        [0].6   // Pylon Home Sensor/Encoder Incongruence - -B26002I -B26007I
        [0].7   // Pylon Home Sensor/Encoder Incongruence - -B26002I -B26007I
        [2].30   // Code 2.30 Pylon Angle overlimit Alarm by Encoder
        [2].16   // Code 2.16 DC Converter Mot 1_3 Rif. T608C DRIVE FAULT
        [0].2   // Gondola Motor 5 Overvoltage Ref. K706C
        [0].10   // Compressor Motor Protection Feedback -F18002C
        [0].0   // Motor 1 Overvoltage control - Relay OK -K10302G
        [1].0   // Gondola Communication Modem Fault CH1 & CH2 -T27002C
        [0].11   // Motor 5 Overvoltage control - Relay OK -K14302G
        [1].1   // Code 1.1 Contactor QC8201H Fault feedback OFF status
        [1].3   // Code 1.3 Contactor QC8204H Fault feedback OFF status
        [0].12   // Motor 6 Overvoltage control - Relay OK -K14307G
        [0].1   // Motor 2 Overvoltage control - Relay OK -K10307G
        [1].5   // Code 1.5 Contactor QC8206H Fault feedback OFF status
        [1].2   // Code 1.2 Contactor QC8201H Fault feedback ON status
        [0].3   // Motor 3 Overvoltage control - Relay OK -K12302G
        [1].4   // Code 1.4 Contactor QC8204H Fault feedback ON status
        [0].4   // Motor 4 Overvoltage control - Relay OK -K12307G
        [1].6   // Code 1.6 Contactor QC8206H Fault feedback ON status
        [1].7   // Pylon Motor 2/4 Fault
        [1].8   // Pylon Motor 1/3 Fault
   Emergencies_Std_CL1 : DINT[8];
        [1].0   // Motor 1-2 Fan Protection Feedback -F10402C -F10406C
        [1].2   // Motor 3-4 Fan Protection Feedback -F12402C -F12406C
        [1].11   // Motor 5 Thermal Probe -K14702H
        [1].3   // Motor 5-6 Fan Protection Feedback -F14402C -F14406C
        [1].12   // Motor 4 Thermal Probe -K12704H
        [1].13   // Motor 6 Thermal Probe -K14704H
        [2].0   // Module K20510C Fault
        [2].1   // Module K20511C Fault
        [2].2   // Module K20512C Fault
        [2].3   // Module K20513C Fault
        [2].4   // Module K20514C Fault
        [2].5   // Module K20515C Fault
        [2].6   // Module K20516C Fault
        [2].7   // Module K20517C Fault
        [1].14   // Motor 7 Thermal Probe -K16602H
        [1].1   // Motor 7 Fan Protection Feedback -F16402C
        [1].6   // MCC High temeprature -S75003C
        [1].8   // Motor 1 Thermal Probe -K10702H
        [1].9   // Motor 2 Thermal Probe -K10704H
        [1].4   // Gondola Motor 7 Fault
        [1].5   // Pylon Motor 5/6 Fault
   Emergency_Brake_manual_Cmd : BOOL;
   Emergency_Brake_manual_Perm : BOOL := 1;
   Emergency_Brake_SL : ALIAS FOR K300_OCC:6:O.6;   // _S31207D
   Emergency_Captr : DINT[11] := ([0] := 1024, [1] := 384, [2] := 1062171331, [4] := 1062171331);
   Enable_to_Start : UDT_CROUT := (CROUT.Feedback1 := 1, CROUT.Feedback2 := 1, CROUT.InputStatus := 1, CROUT.OutputStatus := 1, CROUT.FeedbackReactionTime := 200, Out_Status := 1);   // Abilitazione allo start QC8011E QC8013E
   Encoder_Resetted : BOOL;
   Fault_2_4 : Powerflex_DC_Fault := (Fault_Code := 75);
   Fault_7 : Powerflex_DC_Fault := (Fault_Code := 75);
   FeedBack_Drives_Contactors : BOOL := 1;
   First_Push_Set_Torque_to_Zero : BOOL;
   Flyng_Start_Req : BOOL;
   Gate_Entry_Unlock_Selector : BOOL := 1;   // -S30701F
   Gate_Exit_Unlock_Selector : BOOL := 1;   // -S30705F
   Gate_Magnalock_Enable : UDT_CROUT := (CROUT.Actuate := 1, CROUT.InputStatus := 1, CROUT.OutputStatus := 1, CROUT.FeedbackReactionTime := 250, CROUT.FP := 1, CROUT.FaultCode := 20483);   // Gate Lock Enable -Q25102E
   Gate_Operator_Unlock_Selector : BOOL;   // -S30707F
   GateCommand : DINT := 416;
        .5   // Gate 1 Open
        .7   // Gate 2 Open
        .9   // Gate 3 Open
        .4   // Gate 1 Close
        .6   // Gate 2 Close
        .8   // Gate 3 Close
   GateRequest : DINT;
        .5   // Gate 1 Open
        .7   // Gate 2 Open
        .9   // Gate 3 Open
        .4   // Gate 1 Close
        .6   // Gate 2 Close
        .8   // Gate 3 Close
   Gates_Auto_Release : BOOL;   // .. At end of Cycle Open Gates Open RESTRAINTS
   Gates_Open_Permissive : Permissive := (All_Permissive_Ok := 1, BitsConditions := -1);
   Girella_Field_Actuate_During_Inactivity : BOOL;
   Girella_Gradi_Sec : DINT := 20;
   Gondola_Axe : Axe := (Speed := -5.538001e-24, Speed_ABS := 5.538001e-24);
   Gondola_Decc_timer_Start : BOOL;
   Gondola_Direction_CW_1 : BOOL;   // 0 > CCW 1 > CW
   Gondola_Direction_CW_2 : BOOL := 1;   // 0 > CCW 1 > CW
   Gondola_Drive_Enable : UDT_CROUT := (CROUT.Feedback1 := 1, CROUT.Feedback2 := 1, CROUT.InputStatus := 1, CROUT.OutputStatus := 1, CROUT.FeedbackReactionTime := 1000);   // Gondola Drive Ch1-Ch2 Start Enable Contactors -Q16105E -Q16107E
   Gondola_Immediatly_Stop : BOOL := 1;
   Gondola_Out_Ref : INT;
   Gondola_Speed_Ref_ABS : REAL;
   Gondola_Speed_Reference : DINT;
   Gondola_Standstill_from_inertia : BOOL := 1;
   Gondola_Stop_Beginning : BOOL;
   Gondola_Stop_CW : BOOL := 1;   // Gondola Sto Direction 0 > CCW 1 > CW
   Gondola_Stop_IP : BOOL;   // Gondola Stop Sequence In Progress
   Gondola_Stop_Step : DINT;
   Gondola_Torque_Lim : REAL := 100.0;
   HLL_T1_R011 : HL_LIMIT := (HighLimit := 77.39982, LowLimit := -77.39982);
   HMI_Angle : REAL;
   HMI_Auto_Cycle_in_Modify : Auto_Cycle := (Pylon_Angle := 120, Cycle_Time_min := 2, Cycle_Time_sec := 25, Gondola_Speed[0] := 20, Gondola_Speed[1] := 70, Gondola_Speed[2] := -75, Gondola_Speed[3] := 50, Gondola_Time[1] := 60, Gondola_Time[2] := 50, Gondola_Time[3] := 20);
   HMI_Auto_Cycle_Step_Modify : DINT := 2;
   HMI_button_addtoindex : BOOL;
   HMI_button_subtracttoindex : BOOL;
   HMI_Current_Screen : DINT;
   HMI_Disable_external_acces : BOOL;   // ROUTER A72A07D Disable external acces
   HMI_Drive_Fault_Descr : STRING[4] := ([1] := 'Communication card fault Port 5', [2] := 'Pommunication card fault Port 5', [3] := 'Pommunication card fault Port 5');
        [0]   // Pylon motor 1 3
        [1]   // Pylon motor 2 4
        [2]   // Gondola motor 5
   HMI_Enable_external_acces : BOOL;   // ROUTER A72A07D Eneble external acces
   HMI_Gondola_Start_Delay : DINT := 5;
   HMI_Horn_Pb : BOOL;   // HMIN Horn Pushbutton
   HMI_JM_Stats_Hist : Run_Count_Hist_JM[10];
   HMI_Lamp_Test : BOOL;
   HMI_Light_Pb : BOOL;
   HMI_Modify_Auto_Cycle_Ptr : DINT := 1;
   HMI_Monitor_Bars_Time : DINT := 500;
   HMI_Overspeed_Test_Pb : BOOL;
   HMI_PAGE_PROOF_TEST : DINT := 2000;
   HMI_Pb_Platform_Open : BOOL;   // HMI Platform Open Command
   HMI_Platform_Close : BOOL;   // HMI Platform Close Command
   HMI_Pylon_Start_Delay : DINT;
   HMI_Remote_Display : DINT := 340;   // Display control 0 = operator 0 <> PLC
   HMI_Remote_Status : DINT;   // 0 = Disabled 1 = Enable but not remote control 2 = Remote control active
   HMI_Reset_Encoder_Position : BOOL;
   HMI_Save_Recipe : BOOL;
   HMI_Status_Safety : Status_Safety := (SafetyLockedState := 1, SafetySignatureExists := 1, SafetySignature := 'A43AB79F09EF4071A8C056133A684EE54B2D7E13DC79E37EC57662737DD5528B', Date := '12/01/2025, 06:58:26.072 PM');
   HMI_Step_in_Modify_Gondola_Speed : DINT := -75;
   HMI_Step_in_Modify_Gondola_Time : DINT := 50;
   HMI_Update_Time : BOOL;
   HMI_Work_Auto_Cycle_Ptr : DINT := 2;
   I_ADSL_Fault_Ch1 : BOOL := 1;   // Gondola Communication Modem Fault CH1 -T27002C
   I_ADSL_Fault_Ch2 : BOOL := 1;   // Gondola Communication Modem Fault CH2 -T27002C
   I_Compressor_Min_Pressure : BOOL := 1;   // Line Pressure Switch - Minimum Pressure -S21504B
   I_Compressor_Motor_Protection : BOOL := 1;   // Compressor Motor Protection Feedback -F18002C
   I_Compressor_Work_Pressure : BOOL;   // Line Pressure Switch - Working Pressure -S21502B
   I_Dryer_Motor_Protection : BOOL := 1;   // Dryer Motor Protection Feedback -F18202C
   I_EStop_Pb_OCC1 : UDT_DCI_STOP_TEST := (Push_Botton.ChannelA := 1, Push_Botton.ChannelB := 1, Push_Botton.InputStatus := 1, Push_Botton.TestRequest := 1, Push_Botton.DiscrepancyTime := 500, Push_Botton.O1 := 1, Status := 1, Test_Request := 1);   // +OCC E-stop -S30301F
   I_EStop_Pb_OCC2 : UDT_DCI_STOP_TEST := (Push_Botton.ChannelA := 1, Push_Botton.ChannelB := 1, Push_Botton.InputStatus := 1, Push_Botton.TestRequest := 1, Push_Botton.DiscrepancyTime := 500, Push_Botton.O1 := 1, Status := 1, Test_Request := 1);   // +OCC2 E-Stop -S28502F
   I_Fbk_Platform_Main_Valve : UDT_DCS := (Dual_Chanel_Stop.InputStatus := 1, Dual_Chanel_Stop.RestartType := 1, Dual_Chanel_Stop.ColdStartType := 1, Dual_Chanel_Stop.SafetyFunction := 100, Dual_Chanel_Stop.DiscrepancyTime := 100, Status := 1);   // Feedback Platform Main Valve -B21902I
   I_Fire_Interface : UDT_DCM := (Dual_Chanel_Monitor.InputStatus := 1, Dual_Chanel_Monitor.SafetyFunction := 100, Dual_Chanel_Monitor.DiscrepancyTime := 1000, Dual_Chanel_Monitor.IS := 1, Status := 1);   // Page 44
   I_Gate_1_Opened : BOOL;   // Gate 1 RFID Sensor Closed -B24501J
   I_Gate_2_Opened : BOOL;   // Gate 2 RFID Sensor Closed -B24601J
   I_Gate_3_Opened : BOOL;   // Gate 3 RFID Sensor Closed -B24701J
   I_Gate_4_Opened : BOOL;   // Gate 4 RFID Sensor Closed -B24801J
   I_Gate_DOOR_NEAR_EAC5_Closed : UDT_DCM := (Dual_Chanel_Monitor.InputStatus := 1, Dual_Chanel_Monitor.SafetyFunction := 100, Dual_Chanel_Monitor.DiscrepancyTime := 250, Dual_Chanel_Monitor.IS := 1, Status := 1);   // GATE 4 DOOR NEAR RFID SENSOR - EAC-5 -B24803J
   I_Gate_ENTER_G01_Closed : UDT_DCM := (Dual_Chanel_Monitor.ChannelA := 1, Dual_Chanel_Monitor.ChannelB := 1, Dual_Chanel_Monitor.InputStatus := 1, Dual_Chanel_Monitor.SafetyFunction := 100, Dual_Chanel_Monitor.DiscrepancyTime := 250, Dual_Chanel_Monitor.O1 := 1, Dual_Chanel_Monitor.IS := 1, Status := 1);   // GATE ENTER (G01) -B25204I
   I_Gate_EXIT_G05_Closed : UDT_DCM := (Dual_Chanel_Monitor.ChannelA := 1, Dual_Chanel_Monitor.ChannelB := 1, Dual_Chanel_Monitor.InputStatus := 1, Dual_Chanel_Monitor.SafetyFunction := 100, Dual_Chanel_Monitor.DiscrepancyTime := 250, Dual_Chanel_Monitor.O1 := 1, Dual_Chanel_Monitor.IS := 1, Status := 1);   // GATE EXIT (G05) -B25304I
   I_Gate_OPERATOR_Closed : UDT_DCM := (Dual_Chanel_Monitor.InputStatus := 1, Dual_Chanel_Monitor.SafetyFunction := 100, Dual_Chanel_Monitor.DiscrepancyTime := 250, Dual_Chanel_Monitor.IS := 1, Status := 1);   // GATE 4 OPERATOR RFID SENSOR - MOP -B25404J
   I_Gates_Closed : UDT_DCM := (Dual_Chanel_Monitor.ChannelA := 1, Dual_Chanel_Monitor.ChannelB := 1, Dual_Chanel_Monitor.InputStatus := 1, Dual_Chanel_Monitor.SafetyFunction := 100, Dual_Chanel_Monitor.DiscrepancyTime := 250, Dual_Chanel_Monitor.O1 := 1, Dual_Chanel_Monitor.IS := 1, Status := 1);   // Gate Closed RFID series -B24802J
   I_GMB_RCC1_Temperature_OK : BOOL := 1;   // +GMB_RCC1 Temperature OK -S40103E
   I_Gondola_Home_Position : BOOL := 1;   // Gondola Home Position -B40002I -B40007I
   I_Gondola_Home_Position_Sensor_1 : UDT_DCM := (Dual_Chanel_Monitor.ChannelA := 1, Dual_Chanel_Monitor.InputStatus := 1, Dual_Chanel_Monitor.SafetyFunction := 40, Dual_Chanel_Monitor.InputType := 2, Dual_Chanel_Monitor.DiscrepancyTime := 100, Dual_Chanel_Monitor.O1 := 1, Dual_Chanel_Monitor.IS := 1, Status := 1);   // Home Sensor Speed Check -B40002I
   I_Gondola_Home_Position_Sensor_2 : UDT_DCM := (Dual_Chanel_Monitor.ChannelB := 1, Dual_Chanel_Monitor.InputStatus := 1, Dual_Chanel_Monitor.SafetyFunction := 40, Dual_Chanel_Monitor.InputType := 2, Dual_Chanel_Monitor.DiscrepancyTime := 100, Dual_Chanel_Monitor.IS := 1, Status := 1);   // Home Sensor Speed Check -B40007I
   I_HMI_Login_Enable : BOOL;   // Primary console Key selector Display Login -S30309F
   I_Light_Selector : BOOL := 1;   // Light Selector Switch -S30408F
   I_MCC_Temperature_OK : BOOL := 1;   // MCC temeprature OK -S75003C
   I_Motor_1_2_Fan_Protection_Feedback : BOOL := 1;   // Motor 1-2 Fan Protection Feedback -F10402C -F10406C
   I_Motor_1_Overvoltage_Control : BOOL := 1;   // Motor 1 Overvoltage control - Relay OK -K10302G
   I_Motor_1_Thermal_Probe : BOOL := 1;   // Motor 1 Thermal Probe -K10702H
   I_Motor_2_Overvoltage_Control : BOOL := 1;   // Motor 2 Overvoltage control - Relay OK -K10307G
   I_Motor_2_Thermal_Probe : BOOL := 1;   // Motor 2 Thermal Probe -K10704H
   I_Motor_3_4_Fan_Protection_Feedback : BOOL := 1;   // Motor 3-4 Fan Protection Feedback -F12402C -F12406C
   I_Motor_3_Overvoltage_Control : BOOL := 1;   // Motor 3 Overvoltage control - Relay OK -K12302G
   I_Motor_3_Thermal_Probe : BOOL := 1;   // Motor 3 Thermal Probe -K12702H
   I_Motor_4_Overvoltage_Control : BOOL := 1;   // Motor 4 Overvoltage control - Relay OK -K12307G
   I_Motor_4_Thermal_Probe : BOOL := 1;   // Motor 4 Thermal Probe -K12704H
   I_Motor_5_6_Fan_Protection_Feedback : BOOL := 1;   // Motor 5-6 Fan Protection Feedback -F14402C -F14406C
   I_Motor_5_Overvoltage_Control : BOOL := 1;   // Motor 5 Overvoltage control - Relay OK -K14302G
   I_Motor_5_Thermal_Probe : BOOL := 1;   // Motor 5 Thermal Probe -K14702H
   I_Motor_6_Overvoltage_Control : BOOL := 1;   // Motor 6 Overvoltage control - Relay OK -K14307G
   I_Motor_6_Thermal_Probe : BOOL := 1;   // Motor 6 Thermal Probe -K14704H
   I_Motor_7_Fan_Protection_Feedback : BOOL := 1;   // Motor 7 Fan Protection Feedback -F16402C
   I_Motor_7_Thermal_Probe : BOOL := 1;   // Motor 7 Thermal Probe -K16602H
   I_OCC1_EntGate_PB : BOOL := 1;   // OCC1 Entrance Gate Open/Close -S30701F
   I_OCC1_ExitGate_PB : BOOL := 1;   // OCC1 ExitGate Open/Close -S30707F
   I_OCC1_Stop_Cycle_PB : BOOL := 1;   // Stop Cycle -S30308F
   I_OCC2_ACONFIRM : BOOL;   // OCC2 Allow Main CONFIRM -S28602F
   I_OCC2_Disable : UDT_DCM := (Dual_Chanel_Monitor.InputStatus := 1, Dual_Chanel_Monitor.SafetyFunction := 100, Dual_Chanel_Monitor.DiscrepancyTime := 3000, Dual_Chanel_Monitor.IS := 1, Status := 1);   // OCC 2 CONTROL DISABLE Page 310
   I_OCC2_ExitGate_PB : BOOL;   // OCC2 ExitGate Open/Close -S28507F
   I_OCC2_RESTRAINTS_RELEASE : Sel_3_Pos_2_Input := (Status_Ch_1 := 1, Status_Ch_2 := 1, Center := 1);   // -S28507F RESTRAINTS RELEASE UNLOCK -RUN- LOCK
   I_OCC2_Stop_Cycle_PB : BOOL := 1;   // Stop Cycle -S28606F
   I_OCC_Aut_Man_Selector_Motion : UDT_DCM := (Dual_Chanel_Monitor.ChannelA := 1, Dual_Chanel_Monitor.InputStatus := 1, Dual_Chanel_Monitor.SafetyFunction := 100, Dual_Chanel_Monitor.InputType := 2, Dual_Chanel_Monitor.DiscrepancyTime := 500, Dual_Chanel_Monitor.O1 := 1, Dual_Chanel_Monitor.IS := 1, Status := 1);   // S30801F
   I_OCC_Emergency_Brake : BOOL;   // I OCC Emergency Brake -S31207D
   I_OCC_LockOut_Motion : UDT_DCM := (Dual_Chanel_Monitor.ChannelA := 1, Dual_Chanel_Monitor.ChannelB := 1, Dual_Chanel_Monitor.InputStatus := 1, Dual_Chanel_Monitor.SafetyFunction := 100, Dual_Chanel_Monitor.DiscrepancyTime := 500, Dual_Chanel_Monitor.O1 := 1, Dual_Chanel_Monitor.IS := 1, Status := 1);   // OCC -Lockout Motion -Q31203E
   I_OCC_Memory_Footpedal : BOOL := 1;
   I_OCC_Operator_Enable_Key : BOOL := 1;   // OCC Console Enabled -S30305F
   I_OCC_Temperature_OK : BOOL := 1;   // OCC temperature OK -S31003E
   I_Operator_Footpedal : BOOL := 1;   // Operator Footpedal -S30901F
   I_Platform_Closed : UDT_DCM := (Dual_Chanel_Monitor.ChannelA := 1, Dual_Chanel_Monitor.ChannelB := 1, Dual_Chanel_Monitor.InputStatus := 1, Dual_Chanel_Monitor.SafetyFunction := 41, Dual_Chanel_Monitor.DiscrepancyTime := 200, Dual_Chanel_Monitor.O1 := 1, Dual_Chanel_Monitor.IS := 1, Status := 1);   // Platform Closed RFID Series -B22501J... -B22807J -B22801B
   I_Platform_Line_Min_Pressure_Switch : BOOL;   // Platform Line Minimum Pressure Switch -S21511B
   I_Platform_Line_Unlock_Pressure_Switch : BOOL;   // Unlock Platform Line Pressure Switch -S22006B
   I_Platform_Opened : UDT_DCM := (Dual_Chanel_Monitor.InputStatus := 1, Dual_Chanel_Monitor.SafetyFunction := 41, Dual_Chanel_Monitor.DiscrepancyTime := 20, Dual_Chanel_Monitor.IS := 1, Status := 1);   // Platform Opened RFID Series -Q23801J -Q23807J
   I_Platform_Pressure_on_Close_Circuit : BOOL;   // Platform Maximum Closing Pressure -S21510B
   I_Platform_Pressure_on_Open_Circuit : BOOL := 1;   // Platform Maximum Opening Pressure -S21507B
   I_Pylon_Home_Ch1 : UDT_DCM := (Dual_Chanel_Monitor.ChannelA := 1, Dual_Chanel_Monitor.InputStatus := 1, Dual_Chanel_Monitor.SafetyFunction := 41, Dual_Chanel_Monitor.InputType := 2, Dual_Chanel_Monitor.DiscrepancyTime := 50, Dual_Chanel_Monitor.O1 := 1, Dual_Chanel_Monitor.IS := 1, Status := 1);   // Home position Pylon Ch1 -B26002I
   I_Pylon_Home_Ch2 : UDT_DCM := (Dual_Chanel_Monitor.ChannelA := 1, Dual_Chanel_Monitor.InputStatus := 1, Dual_Chanel_Monitor.SafetyFunction := 41, Dual_Chanel_Monitor.InputType := 2, Dual_Chanel_Monitor.DiscrepancyTime := 50, Dual_Chanel_Monitor.O1 := 1, Dual_Chanel_Monitor.IS := 1, Status := 1);   // Home position Pylon Ch2 -B26007I
   I_Pylon_Overlimit_Right : UDT_DCS := (Dual_Chanel_Stop.ChannelA := 1, Dual_Chanel_Stop.ChannelB := 1, Dual_Chanel_Stop.InputStatus := 1, Dual_Chanel_Stop.ColdStartType := 1, Dual_Chanel_Stop.SafetyFunction := 100, Dual_Chanel_Stop.DiscrepancyTime := 500, Dual_Chanel_Stop.O1 := 1, Status := 1);   // Pylon Overlimit Switchs -A26510I
   I_RCC_GSA_Temperature_OK : BOOL := 1;   // +RCC_GSA Temperature OK -S50110G
   I_RCC_GSB_Temperature_OK : BOOL := 1;   // +RCC_GSB Temperature OK -S52110G
   I_RCC_GSC_Temperature_OK : BOOL := 1;   // +RCC_GSC Temperature OK -S54110G
   I_RCC_GSD_Temperature_OK : BOOL := 1;   // +RCC_GSD Temperature OK -S56110G
   I_RCC_GSE_Temperature_OK : BOOL := 1;   // +RCC_GSE Temperature OK -S58110G
   I_RCC_GSF_Temperature_OK : BOOL := 1;   // +RCC_GSF Temperature OK -S60110G
   I_RCC_GSG_Temperature_OK : BOOL := 1;   // +RCC_GSG Temperature OK -S62110G
   I_RCC_GSH_Temperature_OK : BOOL := 1;   // +RCC_GSH Temperature OK -S64110G
   I_Remote_Connection_Enabled : BOOL := 1;   // Remote Connection active ROUTER eWON K74A04E
   I_RESTRAINTS_Close_Limit_Switch : BOOL := 1;   // Main Valve Close Limit Switch -B40508I
   I_RESTRAINTS_MainValve_Cosed : BOOL := 1;   // Main Valve Close Limit Switch -B40508I
   I_RESTRAINTS_Open_Limit_Switch : BOOL := 1;   // Main Valve Open Limit Switch -B40504I
   I_RESTRAINTS_PressureswitchCompressor : BOOL := 1;   // RESTRAINTS Main Valve Pressure Switch -S40602J
   I_RESTRAINTS_Selector : Sel_3_Pos_2_Input := (Status_Ch_1 := 1, Status_Ch_2 := 1, Center := 1);   // RESTRAINTS Selctor -S30505F Left = Open Right = Close Center = Nothing
   I_Start_PB : Start_AOI := (Status_Ch_1 := 1, Status_Ch_2 := 1, Ready := 1);   // Primary console Strat Push botton Right and Left -S30401F -S30403F
   I_Zero_Set_Sensor : BOOL;   // Zero Set Sensor -B11201A
   Impulsi_per_360_gradi : DINT := 129600;
   Impulsi_per_grado : REAL := 360.0;
   Increase_Torque_Limit_Mem : BOOL;
   index_for_stats_hist : DINT;
   Jerk_Time : REAL := 0.3;   // T1 Region 1
   K_Brake : REAL := 20.0;
   K_Inversion : REAL := -10.0;   // Fattore di Inversione
   K_Inversion_SCRV : REAL := -10.0;
   K_Speed : REAL := 100.0;
   K_Speed_Factor : REAL := 12.121212;
   LapBarsMonitor : LapBars_Monitor[41] := ([1].Sensor_Open_Memory := 1, [1].Status := 1, [2].Sensor_Open_Memory := 1, [2].Status := 1, [3].Sensor_Open_Memory := 1, [3].Status := 1, [4].Sensor_Open_Memory := 1, [4].Status := 1, [5].Sensor_Open_Memory := 1, [5].Status := 1, [6].Sensor_Open_Memory := 1, [6].Status := 1, [7].Sensor_Open_Memory := 1, [7].Status := 1, [8].Sensor_Open_Memory := 1, [8].Status := 1, [9].Sensor_Open_Memory := 1, [9].Status := 1, [10].Sensor_Open_Memory := 1, [10].Status := 1, [11].Sensor_Open_Memory := 1, [11].Status := 1, [12].Sensor_Open_Memory := 1, [12].Status := 1, [13].Sensor_Open_Memory := 1, [13].Status := 1, [14].Sensor_Open_Memory := 1, [14].Status := 1, [15].Sensor_Open_Memory := 1, [15].Status := 1, [16].Sensor_Open_Memory := 1, [16].Status := 1, [17].Sensor_Open_Memory := 1, [17].Status := 1, [18].Sensor_Open_Memory := 1, [18].Status := 1, [19].Sensor_Open_Memory := 1, [19].Status := 1, [20].Sensor_Open_Memory := 1, [20].Status := 1, [21].Sensor_Open_Memory := 1, [21].Status := 1, [22].Sensor_Open_Memory := 1, [22].Status := 1, [23].Sensor_Open_Memory := 1, [23].Status := 1, [24].Sensor_Open_Memory := 1, [24].Status := 1, [25].Sensor_Open_Memory := 1, [25].Status := 1, [26].Sensor_Open_Memory := 1, [26].Status := 1, [27].Sensor_Open_Memory := 1, [27].Status := 1, [28].Sensor_Open_Memory := 1, [28].Status := 1, [29].Sensor_Open_Memory := 1, [29].Status := 1, [30].Sensor_Open_Memory := 1, [30].Status := 1,
        [31].Sensor_Open_Memory := 1, [31].Status := 1, [32].Sensor_Open_Memory := 1, [32].Status := 1, [33].Sensor_Open_Memory := 1, [33].Status := 1, [34].Sensor_Open_Memory := 1, [34].Status := 1, [35].Sensor_Open_Memory := 1, [35].Status := 1, [36].Sensor_Open_Memory := 1, [36].Status := 1, [37].Sensor_Open_Memory := 1, [37].Status := 1, [38].Sensor_Open_Memory := 1, [38].Status := 1, [39].Sensor_Open_Memory := 1, [39].Status := 1, [40].Sensor_Open_Memory := 1, [40].Status := 1); {access Read Only}
   Life_of_Machine : Life_of_Machine := (Life_HH := 1822, Partial_Life_HH := 1822, Working_Cycle_Number_Partial := 1907, Working_Cycle_Number_Total := 1907, Working_HH_Partial := 101, Working_HH_Total := 101, Working_Minutes_Partial := 10);
   LPF_T1_R021 : FILTER_LOW_PASS := (WLag := 15.0, Order := 1, RTSTime := 1, DeltaT := 0.005);
   LPF_WLang_Speed_to_Torq : REAL := 15.0;
   Maintenance_mode : BOOL;   // Ciclo manutenzione per rotazione girella
   Max_Empty_Torque : REAL := 84.0;   // 75
   Max_Full_Torque : REAL := 100.0;   // 85
   Max_Gondola_Speed_RPM : REAL := 6.5;
   Max_Gondola_Speed_RPS : REAL := 0.108333334;
   MAX_HMI_Speed_Value : DINT := 100;
   Max_Reference_Output : DINT := 25000;
   Max_Speed_Reference : DINT := 900;
   MCC_71_03 : BOOL[32] := ([2] := 1, [3] := 1, [4] := 1, [5] := 1, [6] := 1, [13] := 1, [14] := 1, [15] := 1, [16] := 1, [17] := 1, [18] := 1, [20] := 1, [31] := 1);
        [25]   // Limit switch platform 8 Closed B5111E
        [22]   // Limit switch platform 5 Closed B5102E
        [23]   // Limit switch platform 6 Closed B5104E
        [24]   // Limit switch platform 7 Closed B51007E
        [14]   // NC Main Contactor Motor 1_3 Rif. QC8201H
        [2]   // Motor DC1 DC3 Fan Protection QM502B QM506B
        [13]   // Limit switch Platform 1 Opened B5402E
        [7]   // NO Home position Gondola B5912C
        [31]   // Compressor Protection Rif. QM1013E
        [3]   // Motor DC5 Fan Protection Rif. QM510B
        [27]   // Limit switch plataform 2 Closed Rif. B5004E
        [17]   // Limit switch Platform 2 Opened B5404E
        [18]   // Limit switch Platform 3 Opened B5407E
        [26]   // Limit switch plataform 1 Closed Rif. B500E
        [28]   // Limit switch platform 3 Closed Rif. B5007E
        [29]   // Limit switch platform 4 Closed Rif. B5011E
        [6]   // Motor DC2 DC4 Fan Protection QM1002B QM1005B
        [20]   // Limit switch Platform 4 Opened B5411E
        [11]   // Compressor Contactor Fbk QC3103E Rif. 67/12
   Mem_All_Rack_Sensor_OFF : BOOL := 1;
   Mem_RESTRAINTS_closed_Correctly : BOOL := 1;
   Min_Speed_Reference : DINT := -900;
   Min_Torque_to_Maintain_Height_Full_Load : REAL := 15.0;
   Min_Torque_to_Maintain_Height_min_Load : REAL := 15.0;
   MODE : BOOL := 1;   // MODE 0 = AUTO 1 = MANUAL -S30801F
   MUL_T1_R011 : FBD_MATH := (SourceA := -10.0);
   No_Automatic_E_Stop_Cl_0_Request : BOOL := 1;
   No_Automatic_E_Stop_Cl_1_Request : BOOL := 1;
   No_Emergencies_CL0 : BOOL := 1;
   No_Emergencies_CL1 : BOOL := 1;
   No_Sfty : Std_to_Sfty := (Seat_Auxiliary_Ch_Memory := 1, I_Fan_Feedback_NO := 1, RFID_Reset := 1, No_Std_Emergencies_CL0 := 1, No_Std_Emergencies_CL1 := 1, Pylon_min_speed := 1, Gondola_min_Speed := 1, Fbk_MainCotnactor_M1_M3 := 1, Fbk_MainContactor_M2_M4 := 1, I_Gondola_Field_Contactor_Fdbk := 1, I_Gondola_Fuse_Power_Supply := 1, Motors_Temperature_Ok := 1, Low_speed_thold_emergency_brake := 1, UPS_RCC.I_Alarm := 1, UPS_RCC.O_Control := 1, UPS_MCC.I_Alarm := 1, UPS_MCC.O_Control := 1, Main_valve_Time := 10, HMI_Page := 400, Date_Time.Year := 2025, Date_Time.Month := 12, Date_Time.Day := 1, Date_Time.Hour := 19, Date_Time.Minute := 40, Date_Time.Second := 55, Date_Time.Milli_sec := 254030);
        .I_Fan_Feedback_NO   // Fan Feedback NO Pag.94
        .I_Fan_Feedback_NC   // Fan Feedback NC Pag.94
        .Reset_Status   // Status Reset -S30803F
   NO_SFTY_GateClosedSeries : BOOL;   // All Gates Closed and Locked
   No_Sfty_Gondola_SpdFeedback_ABS : DINT;
   NOSFTY_GateClosedSeries : BOOL;
   O_Brake_Pylon_Motor : BOOL := 1;
   O_Close_Gate1 : BOOL;   // Gate 1 OCC2 Operator Close = Mag ON
   O_Close_Gate2 : BOOL;   // Gate 2 Exit Close = Mag ON
   O_Close_Gate3 : BOOL := 1;   // Gate 3 Entrance Close = Mag ON
   O_Close_Gates : BOOL;
   O_Close_Platform : BOOL := 1;
   O_Compressor_Cmd : BOOL := 1;
   O_Enable_Gates_Sensors : BOOL;
   O_Enable_Remote_Connection : BOOL;   // ROUTER A72A07D Eneble external acces
   O_Front_Leg_Light : BOOL := 1;   // Fron leg and front light signal -K3204H
   O_Gate_Enter_Lock : ALIAS FOR K208_MCC:2:O.Pt00Data;   // -B25204I
   O_Gate_Exit_Lock : ALIAS FOR K208_MCC:2:O.Pt01Data;   // -B25304I
   O_Gate_Operator_Lock : ALIAS FOR K208_MCC:2:O.Pt02Data;   // -B25404I
   O_Gondola_Pendolum_Light : BOOL := 1;   // Gondola and pendulum light signal -K3206H
   O_OCC2_Alarms_Lamp : BOOL;
   O_OCC2_Alarms_Noise : BOOL;
   O_OCC_EStop_SL : ALIAS FOR K300_OCC:5:O.7;   // -S30301F EMERGENCY
   O_Open_Platform : BOOL;
   O_Pilots_Valve_Platform : BOOL := 1;
   O_Platform_Main_Valve : BOOL := 1;   // Valvola principale piattaforma B21902I
   O_Platform_MainValve : UDT_CROUT := (CROUT.Actuate := 1, CROUT.InputStatus := 1, CROUT.OutputStatus := 1, CROUT.FeedbackReactionTime := 1000, CROUT.O1 := 1, CROUT.O2 := 1, In_Status := 1);   // Platform main valve B21902I
   O_Rear_Leg_Light : BOOL := 1;   // Rear leg and rear light signal -K3202H
   O_RESTRAINTS_Main_Valve : BOOL;   // Main Valve -B40501I
   O_RESTRAINTS_MainValve : UDT_CROUT := (CROUT.Feedback1 := 1, CROUT.Feedback2 := 1, CROUT.InputStatus := 1, CROUT.OutputStatus := 1, CROUT.FeedbackReactionTime := 1000, In_Status := 1);   // Main Valve -B40501I
   O_RESTRAINTS_Valve_Lift : BOOL;   // Steps 03 04 05
   O_Sl_RESTRAINTS_Close : ALIAS FOR K300_OCC:5:O.3;
   O_Start_Signal_2 : ALIAS FOR K300_OCC:5:O.2;   // -S30401F RIDE START
   ONP : DINT;   // Optional Not Present
   Op_Gate_Delay : TIMER := (PRE := 15000, ACC := 15000, EN := 1, DN := 1);
   OS_Start_Stop_Cycle_Started : BOOL;
   Os_to_CW_CCW : BOOL;
   Oscillation_Error : REAL := 119.95556;
   Oscillation_Phase : BOOL;
   Overspeed_Threshold_millisec : DINT := 9231;
   Overspeed_Threshold_sec : REAL := 9.230769;
   Paltform_Cycle_Abborted_Mem : BOOL;   // Paltform Cycle Abborted by Stop Pb Mem
   Pb_Platform_Stop : BOOL := 1;   // Platform Stop Command -S30608F
   Platform_Close_Cycle : Sequencer := (Index := 31, Step_Timer[0].PRE := 1000, Step_Timer[1].PRE := 100, Step_Timer[2].PRE := 1000, Step_Timer[3].PRE := 250, Step_Timer[7].PRE := 250, Step_Timer[8].PRE := 1000, Step_Timer[10].PRE := 1000, Time_Limit[0].PRE := 2000, Time_Limit[1].PRE := 1000, Time_Limit[2].PRE := 5000, Time_Limit[3].PRE := 1000, Time_Limit[4].PRE := 10000, Time_Limit[5].PRE := 30000, Time_Limit[6].PRE := 5000, Time_Limit[7].PRE := 1000, Time_Limit[9].PRE := 5000, Time_Limit[10].PRE := 10000, Started := 1, Started_OFF_Delay := 1, Step_31 := 1);
        .Step_06   // Lettura Piattaforma Chiusa (B50..E-B51..E) Series
        .Step_08   // Spegnimento Valvole Di Chiusura(QV6505E- QV6510E)
        .Step_09   // Attendo un tempo e spengo la valvola main QV6515E
        .Step_31   // Rilevazione Piattaforme chiuse con ciclo Completato
        .Step_01   // Attesa permesso da valvola manuale(QV6610E)
        .Step_04   // Accendo Valvole Di Chiusura(QV6505E- QV6510E)
        .Step_03   // 3 Lettura Pressione Valvola Main QV6515E
        .Step_05   // Verifica pressostrati(B3114D)
        .Step_10   // Controllo pressostato B6603D
        .Step_02   // Apertura valvola main QV6515E
        .Step_07   // Controllo Azzeramento Pressione (B3113D)
   Platform_Close_Permissive : Permissive := (All_Permissive_Ok := 1, BitsConditions := -1);
   Platform_Close_Permissive_OK : BOOL := 1;
   Platform_Closed_Aux : DINT := 1;
        .1   // Platform closed Sector 1 -B22501J
        .2   // Platform closed Sector 2 -B22507J
        .3   // Platform closed Sector 3 -B22601J
        .4   // Platform closed Sector 4 -B22607J
        .5   // Platform closed Sector 5 -B22701J
        .6   // Platform closed Sector 6 -B22707J
        .7   // Platform closed Sector 7 -B22801J
        .8   // Platform closed Sector 8 -B22807J
   Platform_CloseMain_Valve_Aux_Comand : BOOL := 1;   // Valvola principale piattaforma QV6515E
   Platform_Closing_Cycle_Alarms_Ok : BOOL := 1;
   Platform_Fbk_Valv_Close : BOOL;   // Platform Close Main Valve Limit Switch -B21909I
   Platform_Fbk_Valv_Open : BOOL;   // Platform Open Main Valve Limit Switch -B21905I
   Platform_Manual_Valve : UDT_DCM := (Dual_Chanel_Monitor.SafetyFunction := 41, Dual_Chanel_Monitor.InputType := 2, Dual_Chanel_Monitor.DiscrepancyTime := 250, Dual_Chanel_Monitor.DiagnosticCode := 32);   // Manual Valve Enabling For Platform -B30705B
   Platform_Open_Cycle : Sequencer := (Step_Timer[0].PRE := 1000, Step_Timer[1].PRE := 100, Step_Timer[2].PRE := 1000, Step_Timer[3].PRE := 1000, Step_Timer[4].PRE := 250, Step_Timer[5].PRE := 1000, Step_Timer[6].PRE := 250, Step_Timer[7].PRE := 250, Step_Timer[8].PRE := 250, Step_Timer[9].PRE := 1000, Step_Timer[10].PRE := 1000, Time_Limit[1].PRE := 1000, Time_Limit[2].PRE := 5000, Time_Limit[3].PRE := 1000, Time_Limit[4].PRE := 10000, Time_Limit[5].PRE := 30000, Time_Limit[6].PRE := 5000, Time_Limit[7].PRE := 1000, Time_Limit[8].PRE := 1000, Time_Limit[9].PRE := 5000, Time_Limit[10].PRE := 10000, Time_Limit[31].PRE := 1000, Step_00 := 1);
        .Step_04   // Apertura Valvole Piattaforma(QV6506E-QV6512E)
        .Step_06   // Lettura Piattaforma Aperta (B54..E..B55..E.)
        .Step_11   // Ciclo Apertura Piattaforme Completato, avvio Ciclo giostra
        .Step_08   // Spengo le Valvole di Apertura(QV6506E-QV6512E)
        .Step_Timer[10].DN   // Ciclo Completato
        .Step_10   // Controllo Pressostato(B6603D)
        .Step_05   // Verifica Pressostati(B3113D)
        .Step_03   // Lettura Pressione Pressostato Main(B6603D)
        .Step_07   // Controllo Azzeramento Pressione(B3114D)
        .Step_02   // Apertura Valvola Main(QV6515E)
        .Step_09   // Spengo La Valvola Main(QV6515)
   Platform_Open_Permissive : Permissive := (BitsConditions := -2049);
   Platform_Open_Permissive_Fail_Edge : DINT := -524289;
   Platform_Open_Permissive_Ok : BOOL;
   Platform_Opened_Aux : DINT := 510;
        .1   // Platform Opened Sector 1 -B23501J
        .2   // Platform Opened Sector 2 -B23507J
        .3   // Platform Opened Sector 3 -B23601J
        .4   // Platform Opened Sector 4 -B23607J
        .5   // Platform Opened Sector 5 -B23701J
        .6   // Platform Opened Sector 6 -B23707J
        .7   // Platform Opened Sector 7 -B23801J
        .8   // Platform Opened Sector 8 -B23807J
   Platform_OpenMain_Valve_Aux_Comand : BOOL;   // Valvola principale piattaforma QV6515E
   PltaformClosed_CycleComplete : BOOL := 1;   // Piattaforme chiuse e ciclo completato
   PltaformOpeneded_CycleComplete : BOOL;   // Rilevazione Piattaforme aperte con ciclo Completato
   Power_On_Delay : BOOL := 1;
   Previous_TimeInStation : DINT := 143;
   ProofTest_Req : BOOL;
   pulse_2_sec : TIMER := (PRE := 2000, ACC := 2000, EN := 1, DN := 1);
   PW_Bool : BOOL[32] := ([2] := 1, [3] := 1, [10] := 1);
   PW_Dint : DINT[64] := ([1] := 80, [2] := 120, [3] := -1, [4] := -1, [5] := 4500, [6] := 5500, [7] := 5500, [8] := 10, [9] := -20, [10] := 30, [11] := 100, [12] := 100, [16] := 100, [17] := 100, [18] := 2, [19] := 100, [20] := 10, [21] := 120, [22] := 1, [23] := 4, [24] := 4, [25] := 3, [26] := 4, [27] := 2, [28] := 10, [32] := 1, [34] := 100, [35] := 300);
   Pylon_Axe : Axe := (Position_0_360 := 0.044444446, Position_Sign_180 := 0.044444446, Position_Abs_180 := 0.044444446);
   Pylon_Brake_Motor : UDT_CROUT := (CROUT.Actuate := 1, CROUT.InputStatus := 1, CROUT.OutputStatus := 1, CROUT.FeedbackReactionTime := 500, CROUT.O1 := 1, CROUT.O2 := 1);   // Pylon Brake command -Q10801E
   Pylon_Contactor_OFF : BOOL := 1;
   Pylon_Field_Actuate_During_Inactivity : BOOL;
   Pylon_Filtered_Speed : REAL;
   Pylon_Filtered_Speed_ABS : REAL;
   Pylon_Home_Position : UDT_DCM := (Dual_Chanel_Monitor.ChannelA := 1, Dual_Chanel_Monitor.ChannelB := 1, Dual_Chanel_Monitor.InputStatus := 1, Dual_Chanel_Monitor.SafetyFunction := 41, Dual_Chanel_Monitor.DiscrepancyTime := 3000, Dual_Chanel_Monitor.O1 := 1, Dual_Chanel_Monitor.FP := 1, Dual_Chanel_Monitor.FaultCode := 16386, Status := 1);   // Home position Pylon -B26002I -B26007I
   Pylon_Overspeed_Max_Th : DINT := 101;
   Pylon_Overspeed_min_Th : DINT;
   Pylon_Overspeed_Sensors : DCA_INPUT := (ColdStartType := 1, Tolerance := 50, HighLimit := 101, DiscrepancyTime := 2000, Revision := 1);
   Pylon_Reference : DINT;
   Pylon_Seq_Std : Sequencer_AOI_Std;
   Pylon_Speed : DINT := 92;
   Pylon_Speed_Ref : DINT;
   Pylon_Start_Drive_1_2 : UDT_CROUT := (CROUT.Feedback1 := 1, CROUT.Feedback2 := 1, CROUT.InputStatus := 1, CROUT.OutputStatus := 1, CROUT.FeedbackReactionTime := 500);   // Pylon Start Drive 1 - 2 Contactors -Q9002H -Q9004H -Q10202G
   Pylon_Start_Drive_3_4 : UDT_CROUT := (CROUT.Feedback1 := 1, CROUT.Feedback2 := 1, CROUT.InputStatus := 1, CROUT.OutputStatus := 1, CROUT.FeedbackReactionTime := 500);   // Pylon Start Drive 3 - 4 Contactors -Q9005H -Q9007H -Q12202G
   Pylon_Start_Drive_5_6 : UDT_CROUT := (CROUT.Feedback1 := 1, CROUT.Feedback2 := 1, CROUT.InputStatus := 1, CROUT.OutputStatus := 1, CROUT.FeedbackReactionTime := 500);   // Pylon Start Drive 5 - 6 Contactors -Q9009E -Q9011E4 -Q14202G -Q14202G
   Pylon_Stop_Phase : BOOL;
   Pylon_Stopped_At_Home : BOOL := 1;   // 5s
   Pylon_Torque_Limit : DINT;
   Ratio_HMI_Speed_Ref : REAL := 9.0;
   Real : REAL[32] := ([0] := 0.06436157, [4] := 5.0, [7] := -1.95, [9] := 100.0, [11] := 10.0, [12] := 25.0, [15] := 5.0, [18] := -100.0, [19] := 0.1, [21] := 3.030303);
        [7]   // Test
   Reference_Out_Conversion_Pylon : REAL := 14.619883;
   Reset_Pulse : BOOL;
   Reset_Status_SL_Request : BOOL;
   RESTRAINTS_ChA_Open_Memory : BOOL := 1;
   RESTRAINTS_ChB_Open_Memory : BOOL := 1;
   RESTRAINTS_Closed : BOOL := 1;   // All RESTRAINTS Closed
   RESTRAINTS_Closing : BOOL;
   Restraints_Cycle : Sequencer := (OS[0] := 3, Step_Timer[0].PRE := 2000, Step_Timer[1].PRE := 500, Step_Timer[1].ACC := 520, Step_Timer[1].EN := 1, Step_Timer[1].DN := 1, Step_Timer[2].PRE := 2000, Step_Timer[3].PRE := 2000, Step_Timer[4].PRE := 20000, Step_Timer[5].PRE := 1000, Step_Timer[6].PRE := 1000, Step_Timer[7].PRE := 1500, Step_Timer[7].ACC := 1520, Step_Timer[7].EN := 1, Step_Timer[7].DN := 1, Step_Timer[20].PRE := 1500, Step_Timer[21].PRE := 500, Step_00 := 1);
        .Step_02   // Apertura valvola principale Attendo il tempo limite per il controllo della tenuta valvole sblocco bracci
        .Step_23   // Rack sensors all activated Close sequence compleated
        .Step_05   // Waiting for LapBars to open
        .Step_01   // Apertura valvola principale Attendo il tempo limite per il controllo della tenuta valvole sblocco bracci